REGION Network 5: Transfer Done To T-103
   RUNG wire#powerrail
      Contact( "R-201_Write_TO_Control_DB"."Transfer_To_T-103_Done" )
      Coil( "Control_Read_FROM_R-201_DB"."Transfer_To_T-103_Done" )
   END_RUNG
   // the same network as SCL:
   "Control_Read_FROM_R-201_DB"."Transfer_To_T-103_Done" := "R-201_Write_TO_Control_DB"."Transfer_To_T-103_Done";
END_REGION

REGION Network 6: Tank Wash done
   RUNG wire#powerrail
      Contact( "R-201_Write_TO_Control_DB".TankWash_done )
      Coil( "Control_Read_FROM_R-201_DB".TankWash_done )
   END_RUNG
   // the same network as SCL:
   "Control_Read_FROM_R-201_DB".TankWash_done := "R-201_Write_TO_Control_DB".TankWash_done;
END_REGION

REGION Network 7: Tube Wash Done
   RUNG wire#powerrail
      Contact( "R-201_Write_TO_Control_DB".TubeWash_Done )
      Coil( "Control_Read_FROM_R-201_DB".TubeWash_Done )
   END_RUNG
   // the same network as SCL:
   "Control_Read_FROM_R-201_DB".TubeWash_Done := "R-201_Write_TO_Control_DB".TubeWash_Done;
END_REGION

REGION Network 8: Idle
   RUNG wire#powerrail
      Contact( "R-201_Write_TO_Control_DB".Idle )
      Coil( "Control_Read_FROM_R-201_DB".Idle )
   END_RUNG
   // the same network as SCL:
   "Control_Read_FROM_R-201_DB".Idle := "R-201_Write_TO_Control_DB".Idle;
END_REGION
END_FUNCTION

// folder: State MACHINE/2)Reactors/Reactor R-201/R-201 <---> Control

FUNCTION "R-201_Signals_FROM_Control" : Void   // FC40, LAD
{ S7_Optimized_Access := 'TRUE' }
VERSION : 0.1
BEGIN

REGION Network 1: Start From Reactor Selector.
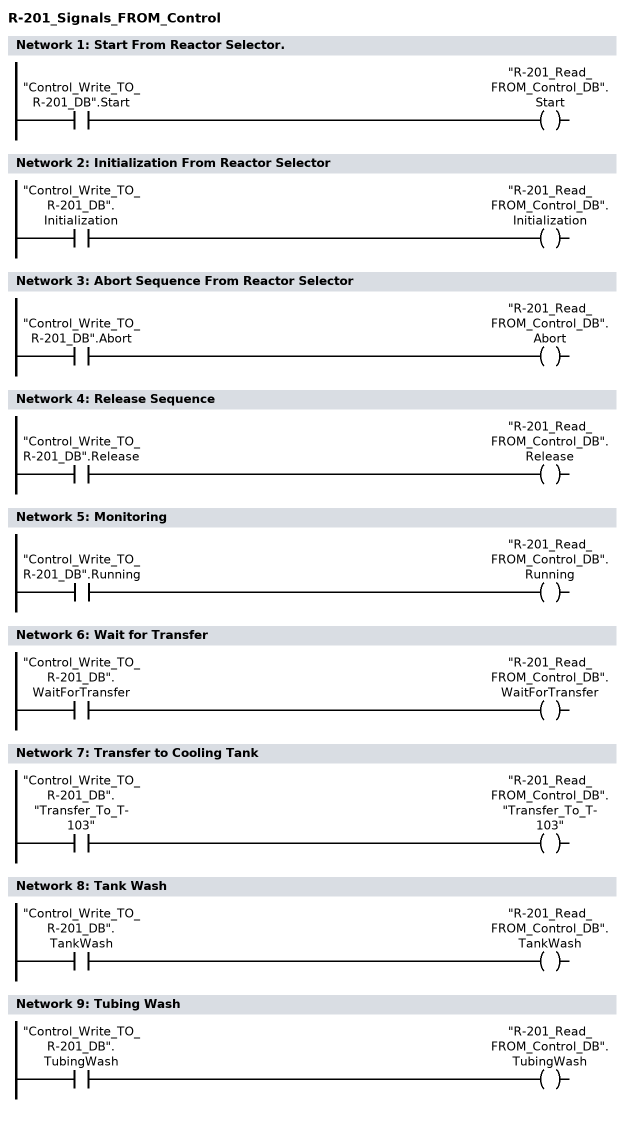
   RUNG wire#powerrail
      Contact( "Control_Write_TO_R-201_DB".Start )
      Coil( "R-201_Read_FROM_Control_DB".Start )
   END_RUNG
   // the same network as SCL:
   "R-201_Read_FROM_Control_DB".Start := "Control_Write_TO_R-201_DB".Start;
END_REGION

REGION Network 2: Initialization From Reactor Selector
   RUNG wire#powerrail
      Contact( "Control_Write_TO_R-201_DB".Initialization )
      Coil( "R-201_Read_FROM_Control_DB".Initialization )
   END_RUNG
   // the same network as SCL:
   "R-201_Read_FROM_Control_DB".Initialization := "Control_Write_TO_R-201_DB".Initialization;
END_REGION

REGION Network 3: Abort Sequence From Reactor Selector
   RUNG wire#powerrail
      Contact( "Control_Write_TO_R-201_DB".Abort )
      Coil( "R-201_Read_FROM_Control_DB".Abort )
   END_RUNG
   // the same network as SCL:
   "R-201_Read_FROM_Control_DB".Abort := "Control_Write_TO_R-201_DB".Abort;
END_REGION

REGION Network 4: Release Sequence
   RUNG wire#powerrail
      Contact( "Control_Write_TO_R-201_DB".Release )
      Coil( "R-201_Read_FROM_Control_DB".Release )
   END_RUNG
   // the same network as SCL:
   "R-201_Read_FROM_Control_DB".Release := "Control_Write_TO_R-201_DB".Release;
END_REGION

REGION Network 5: Monitoring
   RUNG wire#powerrail
      Contact( "Control_Write_TO_R-201_DB".Running )
      Coil( "R-201_Read_FROM_Control_DB".Running )
   END_RUNG
   // the same network as SCL:
   "R-201_Read_FROM_Control_DB".Running := "Control_Write_TO_R-201_DB".Running;
END_REGION

REGION Network 6: Wait for Transfer
   RUNG wire#powerrail
      Contact( "Control_Write_TO_R-201_DB".WaitForTransfer )
      Coil( "R-201_Read_FROM_Control_DB".WaitForTransfer )
   END_RUNG
   // the same network as SCL:
   "R-201_Read_FROM_Control_DB".WaitForTransfer := "Control_Write_TO_R-201_DB".WaitForTransfer;
END_REGION

REGION Network 7: Transfer to Cooling Tank
   RUNG wire#powerrail
      Contact( "Control_Write_TO_R-201_DB"."Transfer_To_T-103" )
      Coil( "R-201_Read_FROM_Control_DB"."Transfer_To_T-103" )
   END_RUNG
   // the same network as SCL:
   "R-201_Read_FROM_Control_DB"."Transfer_To_T-103" := "Control_Write_TO_R-201_DB"."Transfer_To_T-103";
END_REGION

REGION Network 8: Tank Wash
   RUNG wire#powerrail
      Contact( "Control_Write_TO_R-201_DB".TankWash )
      Coil( "R-201_Read_FROM_Control_DB".TankWash )
   END_RUNG
   // the same network as SCL:
   "R-201_Read_FROM_Control_DB".TankWash := "Control_Write_TO_R-201_DB".TankWash;
END_REGION

REGION Network 9: Tubing Wash
   RUNG wire#powerrail
      Contact( "Control_Write_TO_R-201_DB".TubingWash )
      Coil( "R-201_Read_FROM_Control_DB".TubingWash )
   END_RUNG
   // the same network as SCL:
   "R-201_Read_FROM_Control_DB".TubingWash := "Control_Write_TO_R-201_DB".TubingWash;
END_REGION
END_FUNCTION

// folder: State MACHINE/2)Reactors/Reactor R-201/R-201 <---> T-101

FUNCTION "R-201_Signals_FROM_T-101" : Void   // FC61, LAD
{ S7_Optimized_Access := 'TRUE' }
VERSION : 0.1
BEGIN

REGION Network 1: Start Sequence
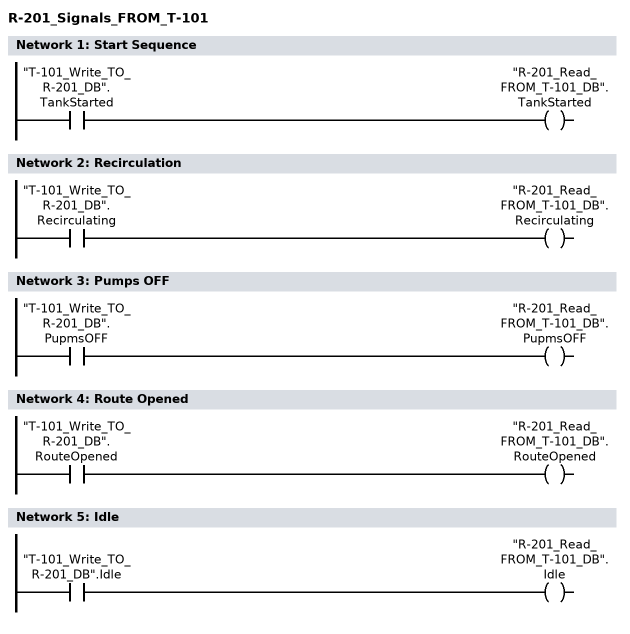
   RUNG wire#powerrail
      Contact( "T-101_Write_TO_R-201_DB".TankStarted )
      Coil( "R-201_Read_FROM_T-101_DB".TankStarted )
   END_RUNG
   // the same network as SCL:
   "R-201_Read_FROM_T-101_DB".TankStarted := "T-101_Write_TO_R-201_DB".TankStarted;
END_REGION

REGION Network 2: Recirculation
   RUNG wire#powerrail
      Contact( "T-101_Write_TO_R-201_DB".Recirculating )
      Coil( "R-201_Read_FROM_T-101_DB".Recirculating )
   END_RUNG
   // the same network as SCL:
   "R-201_Read_FROM_T-101_DB".Recirculating := "T-101_Write_TO_R-201_DB".Recirculating;
END_REGION

REGION Network 3: Pumps OFF
   RUNG wire#powerrail
      Contact( "T-101_Write_TO_R-201_DB".PupmsOFF )
      Coil( "R-201_Read_FROM_T-101_DB".PupmsOFF )
   END_RUNG
   // the same network as SCL:
   "R-201_Read_FROM_T-101_DB".PupmsOFF := "T-101_Write_TO_R-201_DB".PupmsOFF;
END_REGION

REGION Network 4: Route Opened
   RUNG wire#powerrail
      Contact( "T-101_Write_TO_R-201_DB".RouteOpened )
      Coil( "R-201_Read_FROM_T-101_DB".RouteOpened )
   END_RUNG
   // the same network as SCL:
   "R-201_Read_FROM_T-101_DB".RouteOpened := "T-101_Write_TO_R-201_DB".RouteOpened;
END_REGION

REGION Network 5: Idle
   RUNG wire#powerrail
      Contact( "T-101_Write_TO_R-201_DB".Idle )
      Coil( "R-201_Read_FROM_T-101_DB".Idle )
   END_RUNG
   // the same network as SCL:
   "R-201_Read_FROM_T-101_DB".Idle := "T-101_Write_TO_R-201_DB".Idle;
END_REGION
END_FUNCTION

// folder: State MACHINE/2)Reactors/Reactor R-201/R-201 <---> T-102

FUNCTION "R-201_Signals_FROM_T-102" : Void   // FC60, LAD
{ S7_Optimized_Access := 'TRUE' }
VERSION : 0.1
BEGIN

REGION Network 1: Start Sequence
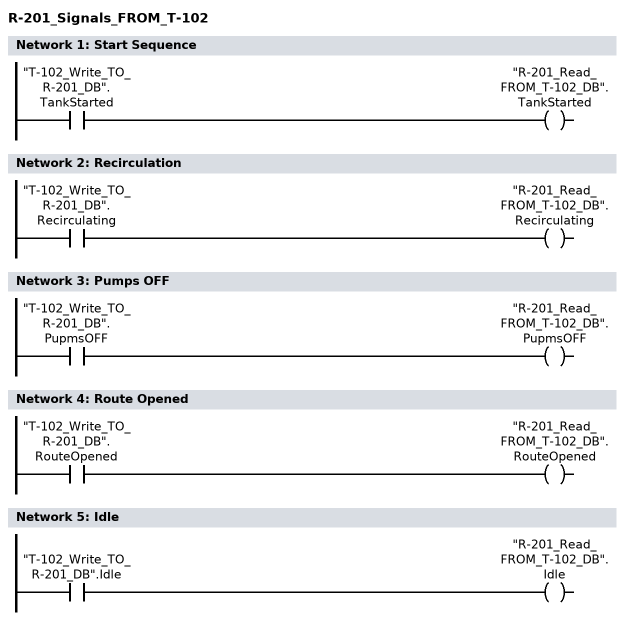
   RUNG wire#powerrail
      Contact( "T-102_Write_TO_R-201_DB".TankStarted )
      Coil( "R-201_Read_FROM_T-102_DB".TankStarted )
   END_RUNG
   // the same network as SCL:
   "R-201_Read_FROM_T-102_DB".TankStarted := "T-102_Write_TO_R-201_DB".TankStarted;
END_REGION

REGION Network 2: Recirculation
   RUNG wire#powerrail
      Contact( "T-102_Write_TO_R-201_DB".Recirculating )
      Coil( "R-201_Read_FROM_T-102_DB".Recirculating )
   END_RUNG
   // the same network as SCL:
   "R-201_Read_FROM_T-102_DB".Recirculating := "T-102_Write_TO_R-201_DB".Recirculating;
END_REGION

REGION Network 3: Pumps OFF
   RUNG wire#powerrail
      Contact( "T-102_Write_TO_R-201_DB".PupmsOFF )
      Coil( "R-201_Read_FROM_T-102_DB".PupmsOFF )
   END_RUNG
   // the same network as SCL:
   "R-201_Read_FROM_T-102_DB".PupmsOFF := "T-102_Write_TO_R-201_DB".PupmsOFF;
END_REGION

REGION Network 4: Route Opened
   RUNG wire#powerrail
      Contact( "T-102_Write_TO_R-201_DB".RouteOpened )
      Coil( "R-201_Read_FROM_T-102_DB".RouteOpened )
   END_RUNG
   // the same network as SCL:
   "R-201_Read_FROM_T-102_DB".RouteOpened := "T-102_Write_TO_R-201_DB".RouteOpened;
END_REGION

REGION Network 5: Idle
   RUNG wire#powerrail
      Contact( "T-102_Write_TO_R-201_DB".Idle )
      Coil( "R-201_Read_FROM_T-102_DB".Idle )
   END_RUNG
   // the same network as SCL:
   "R-201_Read_FROM_T-102_DB".Idle := "T-102_Write_TO_R-201_DB".Idle;
END_REGION
END_FUNCTION

// folder: State MACHINE/2)Reactors/Reactor R-201/R-201 <---> T-103 (CoolingTank)

FUNCTION "R-201_Signals_FROM_T-103" : Void   // FC48, LAD
{ S7_Optimized_Access := 'TRUE' }
VERSION : 0.1
BEGIN

REGION Network 1: Start Sequence
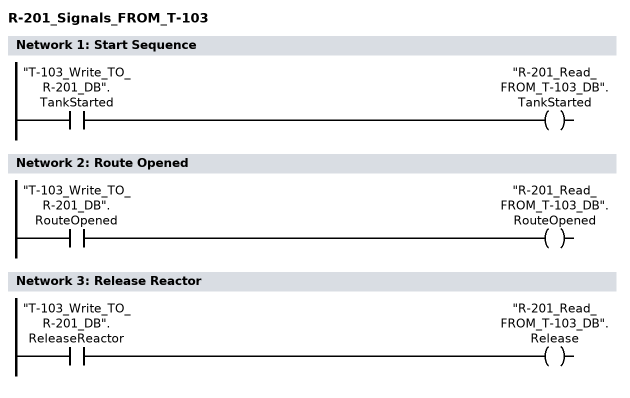
   RUNG wire#powerrail
      Contact( "T-103_Write_TO_R-201_DB".TankStarted )
      Coil( "R-201_Read_FROM_T-103_DB".TankStarted )
   END_RUNG
   // the same network as SCL:
   "R-201_Read_FROM_T-103_DB".TankStarted := "T-103_Write_TO_R-201_DB".TankStarted;
END_REGION

REGION Network 2: Route Opened
   RUNG wire#powerrail
      Contact( "T-103_Write_TO_R-201_DB".RouteOpened )
      Coil( "R-201_Read_FROM_T-103_DB".RouteOpened )
   END_RUNG
   // the same network as SCL:
   "R-201_Read_FROM_T-103_DB".RouteOpened := "T-103_Write_TO_R-201_DB".RouteOpened;
END_REGION

REGION Network 3: Release Reactor
   RUNG wire#powerrail
      Contact( "T-103_Write_TO_R-201_DB".ReleaseReactor )
      Coil( "R-201_Read_FROM_T-103_DB".Release )
   END_RUNG
   // the same network as SCL:
   "R-201_Read_FROM_T-103_DB".Release := "T-103_Write_TO_R-201_DB".ReleaseReactor;
END_REGION
END_FUNCTION

// folder: State MACHINE/2)Reactors/Reactor R-201/R-201 <---> T-104 (WaterSystem)

FUNCTION "R-201_Signals_FROM_T-104" : Void   // FC46, LAD
{ S7_Optimized_Access := 'TRUE' }
VERSION : 0.1
BEGIN

REGION Network 1: Start Sequence
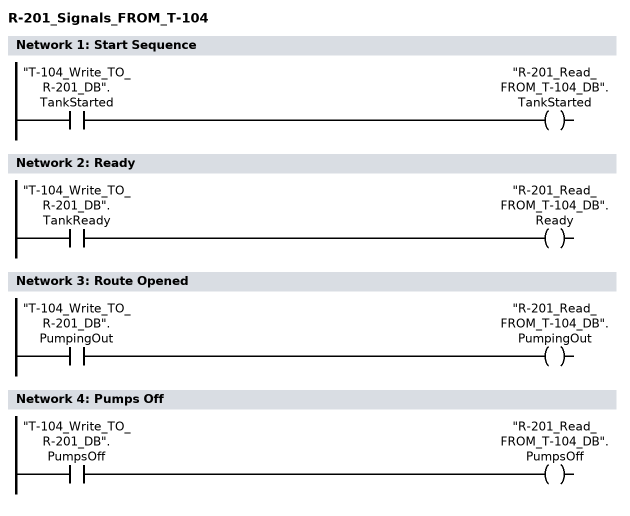
   RUNG wire#powerrail
      Contact( "T-104_Write_TO_R-201_DB".TankStarted )
      Coil( "R-201_Read_FROM_T-104_DB".TankStarted )
   END_RUNG
   // the same network as SCL:
   "R-201_Read_FROM_T-104_DB".TankStarted := "T-104_Write_TO_R-201_DB".TankStarted;
END_REGION

REGION Network 2: Ready
   RUNG wire#powerrail
      Contact( "T-104_Write_TO_R-201_DB".TankReady )
      Coil( "R-201_Read_FROM_T-104_DB".Ready )
   END_RUNG
   // the same network as SCL:
   "R-201_Read_FROM_T-104_DB".Ready := "T-104_Write_TO_R-201_DB".TankReady;
END_REGION

REGION Network 3: Route Opened
   RUNG wire#powerrail
      Contact( "T-104_Write_TO_R-201_DB".PumpingOut )
      Coil( "R-201_Read_FROM_T-104_DB".PumpingOut )
   END_RUNG
   // the same network as SCL:
   "R-201_Read_FROM_T-104_DB".PumpingOut := "T-104_Write_TO_R-201_DB".PumpingOut;
END_REGION

REGION Network 4: Pumps Off
   RUNG wire#powerrail
      Contact( "T-104_Write_TO_R-201_DB".PumpsOff )
      Coil( "R-201_Read_FROM_T-104_DB".PumpsOff )
   END_RUNG
   // the same network as SCL:
   "R-201_Read_FROM_T-104_DB".PumpsOff := "T-104_Write_TO_R-201_DB".PumpsOff;
END_REGION
END_FUNCTION

// folder: State MACHINE/2)Reactors/Reactor R-202

FUNCTION_BLOCK "R-202_SEQ"   // FB34, GRAPH_PLUS
{ S7_Optimized_Access := 'TRUE' }
VERSION : 0.1
   VAR_INPUT
      OFF_SQ : Bool := false;   // Turn sequence off
      INIT_SQ : Bool := false;   // Set sequence to initial state
      ACK_EF : Bool := false;   // Acknowledge all errors and faults
   END_VAR
   VAR_OUTPUT
      S_NO : Int := 0;   // Step number
      S_MORE : Bool := false;   // More steps are available and can be shown in S_NO
      S_ACTIVE : Bool := false;   // Step indicated in S_NO is active
      ERR_FLT : Bool := false;   // Interlock or supervision group error
      AUTO_ON : Bool := false;   // Automatic mode is active
   END_VAR
   VAR
      Reactor : Struct   // Reactor Ctrl
         IDLE : Bool;
         INITIALIZATION : Bool;   // Sequence initialization
         START : Bool;
         DONE_REACTING : Bool;
         COMPLETE : Bool;   // Reactor Complete Read only
         PARA : Bool;   // PARA load Batch side button
         ABORTING : Bool;   // Sequence about
         WAIT : Bool;   // Wating for Permissive read only
      END_STRUCT;
      "Aux Reactor" : Struct
         INITIALIZATION : Bool;
         START : Bool;
         DONE : Bool;
         COMPLETE : Bool;
         PARA : Bool;
         "SELECT_R-203" : Bool;
         "SELECT_R-202" : Bool;
         "SELECT_R-202/R-202" : Bool;
         "SELECT_R-202_T-104" : Bool;
         "SELECT_R-202_T-103" : Bool;
         ABORT : Bool;
         WAIT : Bool;
         LV : Bool;
         FLOW : Bool;
         MIX : Bool;
         "Pre-MIX" : Bool;
         REACTOR : Bool;
         WASH : Bool;
         TUBE : Bool;
         "SEQ_R-203" : Bool;
         "SEQ_R-202" : Bool;
         "SEQ_ R-202 & R-202" : Bool;
         "SEQ_T-103_R-203" : Bool;
         "SEQ_T-103_R-202" : Bool;
         BatchVolume : Real;
         Batchsize : Real;
         batchFlow : Real := 1.0;
         "batchFlow_T-102" : Real;
         BatchPH : Real := 7.0;
         "T-101" : Real;
         BatchTemp : Real := 80.0;
         PM : Bool;
         "TIME" : Struct
            "PRE-MIX" : Time;
            PH_DELAY : Time;
            REACTOR : Time;
            WATCH : Time;
            TUBE : Time;
            CountDown : Struct
               "PRE-MIX" : Time;
               PH_DELAY : Time;
               REACTOR : Time;
               WATCH : Time;
               TUBE : Time;
            END_STRUCT;
         END_STRUCT;
         "TIMER" : Struct
            "PRE-MIX" : IEC_TIMER;
            MIX : IEC_TIMER;
            PH_DELAY : IEC_TIMER;
            REACTOR : IEC_TIMER;
            WASH : IEC_TIMER;
            TUBE : IEC_TIMER;
         END_STRUCT;
      END_STRUCT;
      TEMP : Struct
         TANKS_BATCH : Real;
         "EMPTY_LV_0%" : Real;
         "MIN_LV_20%" : Real;
         "MAX_LV_80%" : Real;
         "BELOW_32%" : Real;
         "Greater_8%" : Real;
         "PRE-ADD" : Real;
         X_SOL_SIZE : Real;
         Y_SOL_SIZE : Real;
         PH_MIN : Real;
         PH_MAX : Real;
         OFFSEt : Struct
            MAX : Real;
            MIN : Real;
         END_STRUCT;
      END_STRUCT;
      COOLING : Struct   // Reactor Ctrl
         IDLE : Bool;
      END_STRUCT;
      HMI_INFO : Array[0..16] of UInt;
      IF_PAR : G7_IfParPlus_V6;
      RT_DATA : G7_RTDataPlus_V6;   // Internal data area
      Abort : G7_TransitionPlus_V6;   // Transition structure
      InitializeR : G7_TransitionPlus_V6;   // Transition structure
      "Fill/Pouring" : G7_TransitionPlus_V6;   // Transition structure
      Re : G7_TransitionPlus_V6;   // Transition structure
      "Fill/Pour" : G7_TransitionPlus_V6;   // Transition structure
      WashT : G7_TransitionPlus_V6;   // Transition structure
      WashTub : G7_TransitionPlus_V6;   // Transition structure
      Std : G7_TransitionPlus_V6;   // Transition structure
      StT : G7_TransitionPlus_V6;   // Transition structure
      WatFll : G7_TransitionPlus_V6;   // Transition structure
      StRW : G7_TransitionPlus_V6;   // Transition structure
      RelT : G7_TransitionPlus_V6;   // Transition structure
      PMix : G7_TransitionPlus_V6;   // Transition structure
      OpR : G7_TransitionPlus_V6;   // Transition structure
      TOT_Done : G7_TransitionPlus_V6;   // Transition structure
      PmpOFF : G7_TransitionPlus_V6;   // Transition structure
      IdleTank : G7_TransitionPlus_V6;   // Transition structure
      TS : G7_TransitionPlus_V6;   // Transition structure
      pHCtl : G7_TransitionPlus_V6;   // Transition structure
      pHCtl2 : G7_TransitionPlus_V6;   // Transition structure
      PmpOFF2 : G7_TransitionPlus_V6;   // Transition structure
      T102_Idle : G7_TransitionPlus_V6;   // Transition structure
      PourD : G7_TransitionPlus_V6;   // Transition structure
      ReacTi : G7_TransitionPlus_V6;   // Transition structure
      ReacD : G7_TransitionPlus_V6;   // Transition structure
      Confirm : G7_TransitionPlus_V6;   // Transition structure
      UserBtch : G7_TransitionPlus_V6;   // Transition structure
      "StT-103" : G7_TransitionPlus_V6;   // Transition structure
      Route_Ok : G7_TransitionPlus_V6;   // Transition structure
      MixDone : G7_TransitionPlus_V6;   // Transition structure
      TimeOut : G7_TransitionPlus_V6;   // Transition structure
      EmptyLv : G7_TransitionPlus_V6;   // Transition structure
      LR : G7_TransitionPlus_V6;   // Transition structure
      DneTransf : G7_TransitionPlus_V6;   // Transition structure
      Trans64 : G7_TransitionPlus_V6;   // Transition structure
      Trans66 : G7_TransitionPlus_V6;   // Transition structure
      TWash : G7_TransitionPlus_V6;   // Transition structure
      STW : G7_TransitionPlus_V6;   // Transition structure
      OpRout : G7_TransitionPlus_V6;   // Transition structure
      TW_RW : G7_TransitionPlus_V6;   // Transition structure
      TW_Vfd : G7_TransitionPlus_V6;   // Transition structure
      Trans87 : G7_TransitionPlus_V6;   // Transition structure
      TW_Wng : G7_TransitionPlus_V6;   // Transition structure
      TW_VfdOf : G7_TransitionPlus_V6;   // Transition structure
      Trans90 : G7_TransitionPlus_V6;   // Transition structure
      DneTnkW : G7_TransitionPlus_V6;   // Transition structure
      TE_SWW : G7_TransitionPlus_V6;   // Transition structure
      TuW : G7_TransitionPlus_V6;   // Transition structure
      STuW : G7_TransitionPlus_V6;   // Transition structure
      Trans103 : G7_TransitionPlus_V6;   // Transition structure
      TuWRW : G7_TransitionPlus_V6;   // Transition structure
      TuWGW : G7_TransitionPlus_V6;   // Transition structure
      TuW_SRW : G7_TransitionPlus_V6;   // Transition structure
      TuW_R : G7_TransitionPlus_V6;   // Transition structure
      Trans108 : G7_TransitionPlus_V6;   // Transition structure
      Trans109 : G7_TransitionPlus_V6;   // Transition structure
      PmpsOn : G7_TransitionPlus_V6;   // Transition structure
      ReEmpty : G7_TransitionPlus_V6;   // Transition structure
      PmpsOff : G7_TransitionPlus_V6;   // Transition structure
      OutleClsd : G7_TransitionPlus_V6;   // Transition structure
      DneTubW : G7_TransitionPlus_V6;   // Transition structure
      Init : G7_TransitionPlus_V6;   // Transition structure
      SAut : G7_TransitionPlus_V6;   // Transition structure
      SIn : G7_TransitionPlus_V6;   // Transition structure
      Initd : G7_TransitionPlus_V6;   // Transition structure
      WaterDn : G7_TransitionPlus_V6;   // Transition structure
      Ab : G7_TransitionPlus_V6;   // Transition structure
      AbortOn : G7_TransitionPlus_V6;   // Transition structure
      DneAbort : G7_TransitionPlus_V6;   // Transition structure
      Idle : G7_StepPlus_V6;   // Step structure
      Ready : G7_StepPlus_V6;   // Step structure
      SelectSeq : G7_StepPlus_V6;   // Step structure
      Started : G7_StepPlus_V6;   // Step structure
      StartTanks : G7_StepPlus_V6;   // Step structure
      FillingUpWater : G7_StepPlus_V6;   // Step structure
      StopReqWaterP : G7_StepPlus_V6;   // Step structure
      ReleaseWTank : G7_StepPlus_V6;   // Step structure
      "Pre-Mix" : G7_StepPlus_V6;   // Step structure
      OpenRoutes : G7_StepPlus_V6;   // Step structure
      X : G7_StepPlus_V6;   // Step structure
      FillDone_T101 : G7_StepPlus_V6;   // Step structure
      Close_T101 : G7_StepPlus_V6;   // Step structure
      "T-101_Done" : G7_StepPlus_V6;   // Step structure
      Y : G7_StepPlus_V6;   // Step structure
      pH_Ctrl1 : G7_StepPlus_V6;   // Step structure
      pH_Ctrl2 : G7_StepPlus_V6;   // Step structure
      FillDone_T102 : G7_StepPlus_V6;   // Step structure
      Close_T102 : G7_StepPlus_V6;   // Step structure
      "T-102_Done" : G7_StepPlus_V6;   // Step structure
      ReactingTime : G7_StepPlus_V6;   // Step structure
      ReactingDone : G7_StepPlus_V6;   // Step structure
      "USER Waiting" : G7_StepPlus_V6;   // Step structure
      "USER BatchP" : G7_StepPlus_V6;   // Step structure
      "Start T-103" : G7_StepPlus_V6;   // Step structure
      "R-202-->T-103" : G7_StepPlus_V6;   // Step structure
      MixToClean : G7_StepPlus_V6;   // Step structure
      LastFlushOut : G7_StepPlus_V6;   // Step structure
      Transfering : G7_StepPlus_V6;   // Step structure
      LastFIllUp : G7_StepPlus_V6;   // Step structure
      FirstFlushOut : G7_StepPlus_V6;   // Step structure
      LastFillUpW : G7_StepPlus_V6;   // Step structure
      LastTransfer : G7_StepPlus_V6;   // Step structure
      Done_Transfer : G7_StepPlus_V6;   // Step structure
      Idle_TWash : G7_StepPlus_V6;   // Step structure
      Start_TWash : G7_StepPlus_V6;   // Step structure
      OpenRoute : G7_StepPlus_V6;   // Step structure
      ReqWaterWash : G7_StepPlus_V6;   // Step structure
      "2011 VFD ON & PID AUTO/Wait for 80%_R-202" : G7_StepPlus_V6;   // Step structure
      StopWaterWash : G7_StepPlus_V6;   // Step structure
      "XV-1044_CC_02_R-202" : G7_StepPlus_V6;   // Step structure
      Washing : G7_StepPlus_V6;   // Step structure
      "2011VFD OFF & PID MAN_R-202" : G7_StepPlus_V6;   // Step structure
      USER_MAN_DRAIN : G7_StepPlus_V6;   // Step structure
      Done_TWash : G7_StepPlus_V6;   // Step structure
      Idle_TubWash : G7_StepPlus_V6;   // Step structure
      Start_TubWash : G7_StepPlus_V6;   // Step structure
      "XV-1044_CO_03_R-202" : G7_StepPlus_V6;   // Step structure
      ReqWaterTuW : G7_StepPlus_V6;   // Step structure
      GettingWater : G7_StepPlus_V6;   // Step structure
      StopRqWaterTuW : G7_StepPlus_V6;   // Step structure
      "ReleaseT-104" : G7_StepPlus_V6;   // Step structure
      "XV-1044_CC_03_R-529" : G7_StepPlus_V6;   // Step structure
      "XV-2023_CO_XV-1044_Cc_R-202" : G7_StepPlus_V6;   // Step structure
      "P-202A/B_ON_R-202" : G7_StepPlus_V6;   // Step structure
      Emptying : G7_StepPlus_V6;   // Step structure
      "P-202A/B_OFF_R-202" : G7_StepPlus_V6;   // Step structure
      Close_Outlet : G7_StepPlus_V6;   // Step structure
      Done_TubWash : G7_StepPlus_V6;   // Step structure
      Initialize : G7_StepPlus_V6;   // Step structure
      SetAuto : G7_StepPlus_V6;   // Step structure
      SetInitial : G7_StepPlus_V6;   // Step structure
      Initialized : G7_StepPlus_V6;   // Step structure
      AbortStarting : G7_StepPlus_V6;   // Step structure
      Aborting : G7_StepPlus_V6;   // Step structure
      Abort_Done : G7_StepPlus_V6;   // Step structure
      SINI : Array[0..9] of USInt;
      LSTT : Array[0..68] of USInt;
      ATAJ : Array[0..68] of USInt;
      ATAB : Array[0..68] of USInt;
      PSTT : Array[0..68] of USInt;
      NSTT : Array[0..68] of USInt;
      ASSJ : Array[0..65] of USInt;
      ASSB : Array[0..65] of USInt;
      PTTS : Array[0..65] of USInt;
      NTTS : Array[0..65] of USInt;
      SW_SQTS : Array[0..65] of USInt;
      SWITCH : Array[0..15] of USInt;
      TVX : Array[0..15] of USInt;
      TTX : Array[0..15] of USInt;
      TSX : Array[0..9] of USInt;
      S00X : Array[0..9] of USInt;
      SOFFX : Array[0..9] of USInt;
      SONX : Array[0..9] of USInt;
      SAX : Array[0..9] of USInt;
      SERRX : Array[0..66] of USInt;
      SMX : Array[0..66] of USInt;
      S0X : Array[0..66] of USInt;
      S1X : Array[0..66] of USInt;
      IL_ALARM_INST : Diag_Alarm;
      SUP_ALARM_INST : Diag_Alarm;
      STEP_TIME_ALARM_INST : Diag_Alarm;
      IEC_TIMER_INST : IEC_TIMER;
      TRANSACTION_FLAG : Bool := false;
   END_VAR
   VAR CONSTANT
      "Single R-202 T-101 seq done" : Int := 214;
      "Single R-202 T-102 seq done" : Int := 218;
   END_VAR
   // SINI[0] := 2;
   // LSTT[0] := 63;
   // NSTT[0] := 63;
   // PTTS[0] := 255;
   // TVX[0] := 16#1;
   // TTX[0] := 16#1;
   // TSX[0] := 16#1;
   // S00X[0] := 16#1;
   // SOFFX[0] := 16#1;
   // SONX[0] := 16#1;
   // SAX[0] := 16#1;
   // SERRX[0] := 16#1;
   // SMX[0] := 16#1;
   // S0X[0] := 16#1;
   // S1X[0] := 16#1;
   // LSTT[38] := 255;
   // SINI[3] := 255;
   // LSTT[1] := 59;
   // LSTT[2] := 255;
   // LSTT[3] := 255;
   // LSTT[4] := 3;
   // LSTT[5] := 34;
   // LSTT[6] := 45;
   // LSTT[7] := 255;
   // LSTT[8] := 255;
   // LSTT[9] := 255;
   // LSTT[10] := 255;
   // LSTT[11] := 255;
   // LSTT[12] := 255;
   // LSTT[13] := 255;
   // LSTT[14] := 255;
   // LSTT[15] := 255;
   // LSTT[16] := 255;
   // LSTT[17] := 255;
   // LSTT[18] := 255;
   // LSTT[19] := 255;
   // LSTT[20] := 255;
   // LSTT[21] := 255;
   // LSTT[22] := 255;
   // LSTT[23] := 255;
   // LSTT[24] := 255;
   // LSTT[56] := 255;
   // LSTT[27] := 255;
   // LSTT[57] := 255;
   // LSTT[29] := 255;
   // LSTT[30] := 255;
   // LSTT[31] := 255;
   // LSTT[32] := 255;
   // LSTT[55] := 255;
   // LSTT[62] := 255;
   // LSTT[44] := 255;
   // LSTT[36] := 255;
   // LSTT[66] := 255;
   // LSTT[39] := 255;
   // LSTT[40] := 255;
   // LSTT[41] := 255;
   // LSTT[42] := 255;
   // LSTT[59] := 255;
   // LSTT[58] := 255;
   // LSTT[46] := 255;
   // LSTT[47] := 255;
   // LSTT[50] := 255;
   // LSTT[51] := 255;
   // LSTT[52] := 255;
   // LSTT[53] := 255;
   // LSTT[54] := 255;
   // NSTT[28] := 28;
   // NSTT[65] := 33;
   // ATAJ[1] := 1;
   // ATAJ[2] := 2;
   // ATAJ[3] := 3;
   // ATAJ[4] := 4;
   // ATAJ[5] := 5;
   // ATAJ[6] := 6;
   // ATAJ[7] := 7;
   // ATAJ[8] := 8;
   // ATAJ[9] := 9;
   // ATAJ[10] := 10;
   // ATAJ[11] := 11;
   // ATAJ[12] := 12;
   // ATAJ[13] := 13;
   // ATAJ[14] := 14;
   // ATAJ[15] := 15;
   // ATAJ[16] := 16;
   // ATAJ[17] := 17;
   // ATAJ[18] := 18;
   // ATAJ[19] := 19;
   // ATAJ[20] := 20;
   // ATAJ[21] := 21;
   // ATAJ[22] := 22;
   // ATAJ[23] := 23;
   // ATAJ[24] := 24;
   // ATAJ[25] := 25;
   // ATAJ[26] := 26;
   // ATAJ[27] := 27;
   // ATAJ[28] := 28;
   // ATAJ[29] := 29;
   // ATAJ[30] := 30;
   // ATAJ[31] := 31;
   // ATAJ[32] := 32;
   // ATAJ[33] := 33;
   // ATAJ[34] := 34;
   // ATAJ[35] := 35;
   // ATAJ[36] := 36;
   // ATAJ[37] := 37;
   // ATAJ[38] := 38;
   // ATAJ[39] := 39;
   // ATAJ[40] := 40;
   // ATAJ[41] := 41;
   // ATAJ[42] := 42;
   // ATAJ[43] := 43;
   // ATAJ[44] := 44;
   // ATAJ[45] := 45;
   // ATAJ[46] := 46;
   // ATAJ[47] := 47;
   // ATAJ[48] := 48;
   // ATAJ[49] := 49;
   // ATAJ[50] := 50;
   // ATAJ[51] := 51;
   // ATAJ[52] := 52;
   // ATAJ[53] := 53;
   // ATAJ[54] := 54;
   // ATAJ[55] := 55;
   // ATAJ[56] := 56;
   // ATAJ[57] := 57;
   // ATAJ[58] := 58;
   // ATAJ[59] := 59;
   // ATAJ[60] := 60;
   // ATAJ[61] := 61;
   // ATAJ[62] := 62;
   // ATAJ[63] := 63;
   // ATAJ[64] := 64;
   // ATAJ[65] := 65;
   // ATAB[1] := 2;
   // ATAB[24] := 24;
   // ATAB[3] := 3;
   // ATAB[4] := 5;
   // ATAB[5] := 6;
   // ATAB[6] := 4;
   // ATAB[7] := 7;
   // ATAB[8] := 8;
   // ATAB[9] := 9;
   // ATAB[10] := 10;
   // ATAB[11] := 11;
   // ATAB[12] := 12;
   // ATAB[13] := 13;
   // ATAB[14] := 14;
   // ATAB[15] := 15;
   // ATAB[16] := 16;
   // ATAB[17] := 17;
   // ATAB[18] := 18;
   // ATAB[21] := 21;
   // ATAB[22] := 22;
   // ATAB[23] := 23;
   // ATAB[29] := 29;
   // ATAB[25] := 25;
   // ATAB[26] := 26;
   // ATAB[27] := 27;
   // ATAB[28] := 28;
   // ATAB[30] := 30;
   // ATAB[31] := 31;
   // ATAB[32] := 32;
   // ATAB[33] := 33;
   // ATAB[34] := 34;
   // ATAB[35] := 35;
   // ATAB[36] := 36;
   // ATAB[37] := 37;
   // ATAB[38] := 38;
   // ATAB[39] := 39;
   // ATAB[40] := 40;
   // ATAB[41] := 41;
   // ATAB[42] := 42;
   // ATAB[43] := 43;
   // ATAB[44] := 44;
   // ATAB[45] := 45;
   // ATAB[46] := 46;
   // ATAB[47] := 47;
   // ATAB[48] := 48;
   // ATAB[49] := 49;
   // ATAB[50] := 50;
   // ATAB[51] := 51;
   // ATAB[52] := 52;
   // ATAB[53] := 53;
   // ATAB[54] := 54;
   // ATAB[55] := 55;
   // ATAB[56] := 56;
   // ATAB[57] := 57;
   // ATAB[58] := 58;
   // ATAB[59] := 59;
   // ATAB[60] := 60;
   // ATAB[61] := 61;
   // ATAB[62] := 62;
   // ATAB[63] := 63;
   // ATAB[64] := 64;
   // ATAB[65] := 65;
   // PSTT[33] := 31;
   // PSTT[16] := 12;
   // PSTT[3] := 1;
   // PSTT[4] := 2;
   // PSTT[5] := 2;
   // PSTT[6] := 2;
   // PSTT[7] := 3;
   // PSTT[8] := 4;
   // PSTT[9] := 5;
   // PSTT[10] := 6;
   // PSTT[12] := 8;
   // PSTT[13] := 9;
   // PSTT[60] := 58;
   // PSTT[14] := 10;
   // PSTT[17] := 14;
   // PSTT[18] := 15;
   // PSTT[19] := 16;
   // PSTT[20] := 17;
   // PSTT[21] := 18;
   // PSTT[22] := 13;
   // PSTT[23] := 20;
   // PSTT[24] := 21;
   // PSTT[25] := 22;
   // PSTT[26] := 23;
   // PSTT[27] := 24;
   // PSTT[28] := 25;
   // PSTT[29] := 26;
   // PSTT[30] := 27;
   // PSTT[31] := 28;
   // PSTT[32] := 30;
   // PSTT[40] := 38;
   // PSTT[38] := 36;
   // PSTT[35] := 33;
   // PSTT[36] := 34;
   // PSTT[37] := 35;
   // PSTT[59] := 57;
   // PSTT[41] := 40;
   // PSTT[58] := 56;
   // PSTT[42] := 41;
   // PSTT[43] := 42;
   // PSTT[44] := 43;
   // PSTT[45] := 44;
   // PSTT[46] := 39;
   // PSTT[47] := 45;
   // PSTT[48] := 46;
   // PSTT[49] := 47;
   // PSTT[50] := 48;
   // PSTT[51] := 49;
   // PSTT[52] := 50;
   // PSTT[56] := 54;
   // PSTT[57] := 55;
   // PSTT[61] := 59;
   // PSTT[62] := 60;
   // PSTT[63] := 61;
   // PSTT[64] := 62;
   // PSTT[65] := 29;
   // NSTT[1] := 59;
   // NSTT[2] := 1;
   // NSTT[3] := 2;
   // NSTT[4] := 3;
   // NSTT[5] := 34;
   // NSTT[6] := 45;
   // NSTT[7] := 23;
   // NSTT[8] := 5;
   // NSTT[9] := 6;
   // NSTT[10] := 7;
   // NSTT[11] := 8;
   // NSTT[12] := 9;
   // NSTT[13] := 10;
   // NSTT[14] := 11;
   // NSTT[15] := 12;
   // NSTT[16] := 13;
   // NSTT[17] := 15;
   // NSTT[18] := 16;
   // NSTT[19] := 17;
   // NSTT[20] := 18;
   // NSTT[21] := 19;
   // NSTT[22] := 20;
   // NSTT[23] := 21;
   // NSTT[24] := 22;
   // NSTT[56] := 55;
   // NSTT[27] := 25;
   // NSTT[57] := 56;
   // NSTT[29] := 32;
   // NSTT[30] := 29;
   // NSTT[31] := 30;
   // NSTT[32] := 31;
   // NSTT[55] := 54;
   // NSTT[62] := 61;
   // NSTT[44] := 44;
   // NSTT[36] := 35;
   // NSTT[66] := 64;
   // NSTT[39] := 38;
   // NSTT[40] := 39;
   // NSTT[41] := 41;
   // NSTT[42] := 42;
   // NSTT[59] := 58;
   // NSTT[58] := 57;
   // NSTT[46] := 40;
   // NSTT[47] := 46;
   // NSTT[50] := 49;
   // NSTT[51] := 50;
   // NSTT[52] := 51;
   // NSTT[53] := 52;
   // NSTT[54] := 53;
   // LSTT[65] := 255;
   // ASSJ[1] := 1;
   // ASSJ[2] := 2;
   // ASSJ[3] := 3;
   // ASSJ[4] := 4;
   // ASSJ[5] := 5;
   // ASSJ[6] := 6;
   // ASSJ[7] := 7;
   // ASSJ[8] := 8;
   // ASSJ[9] := 9;
   // ASSJ[10] := 10;
   // ASSJ[11] := 11;
   // ASSJ[12] := 12;
   // ASSJ[13] := 19;
   // ASSJ[14] := 14;
   // ASSJ[15] := 15;
   // ASSJ[16] := 16;
   // ASSJ[17] := 17;
   // ASSJ[18] := 18;
   // ASSJ[19] := 13;
   // ASSJ[20] := 20;
   // ASSJ[21] := 21;
   // ASSJ[22] := 22;
   // ASSJ[23] := 23;
   // ASSJ[24] := 24;
   // ASSJ[25] := 25;
   // ASSJ[26] := 26;
   // ASSJ[27] := 27;
   // ASSJ[28] := 28;
   // ASSJ[29] := 29;
   // ASSJ[30] := 30;
   // ASSJ[31] := 31;
   // ASSJ[32] := 32;
   // ASSJ[33] := 33;
   // ASSJ[34] := 34;
   // ASSJ[35] := 35;
   // ASSJ[36] := 36;
   // ASSJ[37] := 37;
   // ASSJ[38] := 38;
   // ASSJ[39] := 39;
   // ASSJ[40] := 40;
   // ASSJ[41] := 41;
   // ASSJ[42] := 42;
   // ASSJ[43] := 43;
   // ASSJ[44] := 44;
   // ASSJ[45] := 45;
   // ASSJ[46] := 46;
   // ASSJ[47] := 47;
   // ASSJ[48] := 48;
   // ASSJ[49] := 49;
   // ASSJ[50] := 50;
   // ASSJ[51] := 51;
   // ASSJ[52] := 52;
   // ASSJ[53] := 53;
   // ASSJ[54] := 54;
   // ASSJ[55] := 55;
   // ASSJ[56] := 56;
   // ASSJ[57] := 57;
   // ASSJ[58] := 58;
   // ASSJ[59] := 59;
   // ASSJ[60] := 60;
   // ASSJ[61] := 61;
   // ASSJ[62] := 62;
   // ASSJ[63] := 63;
   // ASSB[1] := 1;
   // ASSB[2] := 2;
   // ASSB[3] := 3;
   // ASSB[4] := 4;
   // ASSB[5] := 5;
   // ASSB[6] := 6;
   // ASSB[7] := 7;
   // ASSB[8] := 8;
   // ASSB[9] := 9;
   // ASSB[10] := 14;
   // ASSB[11] := 11;
   // ASSB[12] := 12;
   // ASSB[13] := 13;
   // ASSB[14] := 10;
   // ASSB[15] := 15;
   // ASSB[16] := 16;
   // ASSB[17] := 17;
   // ASSB[18] := 18;
   // ASSB[19] := 19;
   // ASSB[20] := 20;
   // ASSB[21] := 21;
   // ASSB[22] := 22;
   // ASSB[23] := 23;
   // ASSB[24] := 24;
   // ASSB[25] := 25;
   // ASSB[26] := 26;
   // ASSB[27] := 27;
   // ASSB[28] := 28;
   // ASSB[29] := 29;
   // ASSB[30] := 30;
   // ASSB[31] := 31;
   // ASSB[32] := 32;
   // ASSB[33] := 33;
   // ASSB[34] := 34;
   // ASSB[35] := 35;
   // ASSB[36] := 36;
   // ASSB[37] := 37;
   // ASSB[38] := 38;
   // ASSB[39] := 39;
   // ASSB[40] := 40;
   // ASSB[41] := 41;
   // ASSB[42] := 42;
   // ASSB[43] := 43;
   // ASSB[44] := 44;
   // ASSB[45] := 45;
   // ASSB[46] := 46;
   // ASSB[47] := 47;
   // ASSB[48] := 48;
   // ASSB[49] := 49;
   // ASSB[50] := 50;
   // ASSB[51] := 51;
   // ASSB[52] := 52;
   // ASSB[53] := 53;
   // ASSB[54] := 54;
   // ASSB[55] := 55;
   // ASSB[56] := 56;
   // ASSB[57] := 57;
   // ASSB[58] := 58;
   // ASSB[59] := 59;
   // ASSB[60] := 60;
   // ASSB[61] := 61;
   // ASSB[62] := 62;
   // ASSB[63] := 63;
   // PTTS[3] := 255;
   // PTTS[61] := 62;
   // PTTS[5] := 8;
   // PTTS[6] := 9;
   // PTTS[7] := 10;
   // PTTS[8] := 11;
   // PTTS[9] := 12;
   // PTTS[10] := 13;
   // PTTS[11] := 14;
   // PTTS[12] := 15;
   // PTTS[13] := 16;
   // PTTS[14] := 13;
   // PTTS[15] := 17;
   // PTTS[16] := 18;
   // PTTS[17] := 19;
   // PTTS[18] := 20;
   // PTTS[19] := 21;
   // PTTS[20] := 22;
   // PTTS[21] := 23;
   // PTTS[22] := 24;
   // PTTS[23] := 7;
   // PTTS[24] := 255;
   // PTTS[25] := 27;
   // PTTS[26] := 33;
   // SW_SQTS[3] := 2;
   // PTTS[31] := 32;
   // PTTS[32] := 29;
   // PTTS[33] := 65;
   // PTTS[34] := 255;
   // PTTS[35] := 36;
   // PTTS[36] := 37;
   // PTTS[37] := 38;
   // PTTS[38] := 39;
   // PTTS[39] := 40;
   // PTTS[40] := 46;
   // PTTS[41] := 41;
   // PTTS[42] := 42;
   // PTTS[43] := 43;
   // PTTS[44] := 44;
   // PTTS[45] := 255;
   // PTTS[46] := 47;
   // PTTS[47] := 48;
   // PTTS[48] := 49;
   // PTTS[49] := 50;
   // PTTS[50] := 51;
   // PTTS[51] := 52;
   // PTTS[52] := 53;
   // PTTS[53] := 54;
   // PTTS[54] := 55;
   // PTTS[55] := 56;
   // PTTS[56] := 57;
   // PTTS[57] := 58;
   // PTTS[58] := 59;
   // PTTS[59] := 255;
   // PTTS[60] := 61;
   // SW_SQTS[34] := 7;
   // PTTS[62] := 63;
   // PTTS[63] := 255;
   // SW_SQTS[35] := 7;
   // NTTS[3] := 7;
   // NTTS[5] := 9;
   // NTTS[6] := 10;
   // NTTS[7] := 11;
   // NTTS[8] := 12;
   // NTTS[9] := 13;
   // NTTS[10] := 14;
   // NTTS[11] := 15;
   // NTTS[12] := 16;
   // NTTS[13] := 22;
   // NTTS[14] := 17;
   // NTTS[15] := 18;
   // NTTS[16] := 19;
   // NTTS[17] := 20;
   // NTTS[18] := 21;
   // NTTS[19] := 22;
   // NTTS[20] := 23;
   // NTTS[21] := 24;
   // NTTS[22] := 25;
   // NTTS[23] := 26;
   // NTTS[24] := 27;
   // NTTS[25] := 28;
   // NTTS[26] := 29;
   // NTTS[27] := 30;
   // NTTS[28] := 31;
   // NTTS[29] := 65;
   // NTTS[30] := 32;
   // NTTS[31] := 33;
   // NTTS[32] := 34;
   // NTTS[33] := 35;
   // NTTS[34] := 36;
   // NTTS[35] := 37;
   // NTTS[36] := 38;
   // NTTS[37] := 39;
   // NTTS[38] := 40;
   // NTTS[39] := 46;
   // NTTS[40] := 41;
   // NTTS[41] := 42;
   // NTTS[42] := 43;
   // NTTS[43] := 44;
   // NTTS[44] := 45;
   // NTTS[45] := 47;
   // NTTS[46] := 48;
   // NTTS[47] := 49;
   // NTTS[48] := 50;
   // NTTS[49] := 51;
   // NTTS[50] := 52;
   // NTTS[51] := 53;
   // NTTS[52] := 54;
   // NTTS[53] := 55;
   // NTTS[54] := 56;